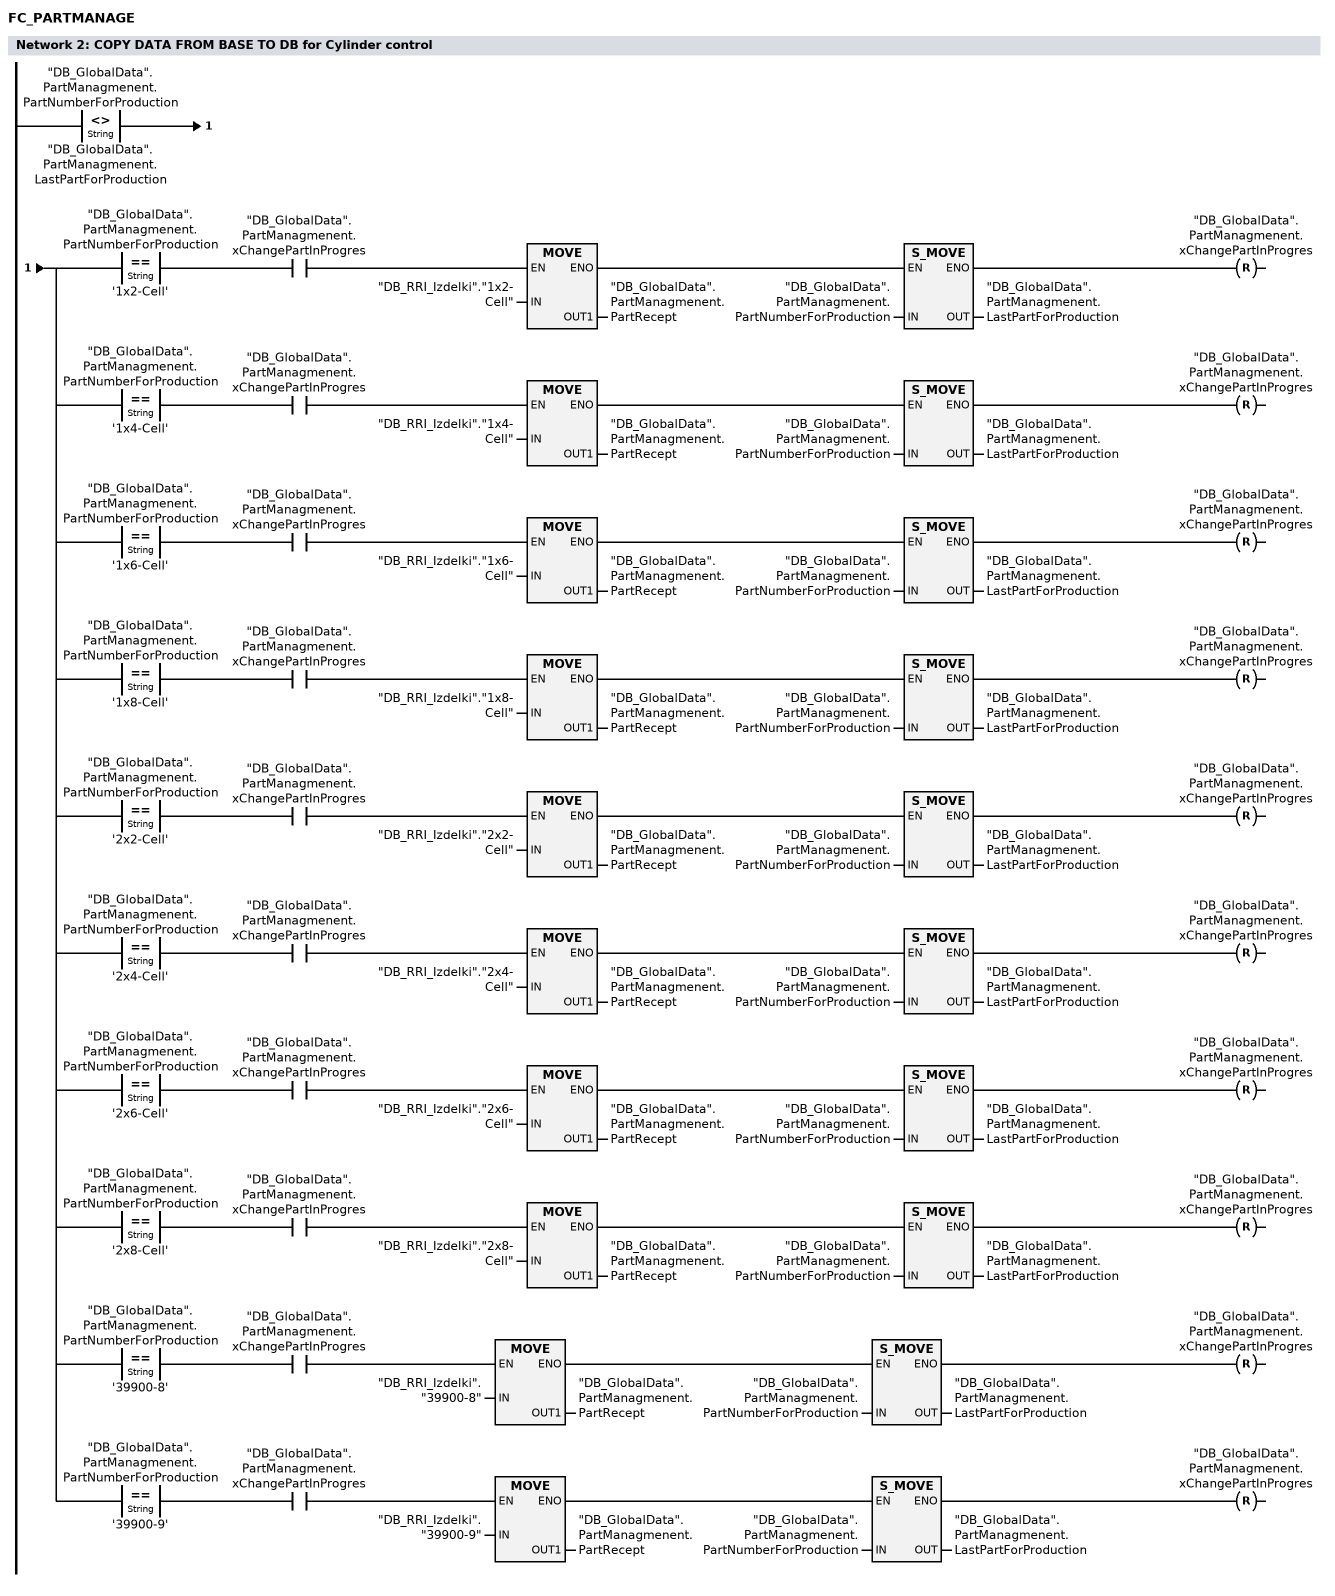
   RUNG wire#powerrail
      { S7_Templates := "SrcType := String" } NE_Contact(in1 := "DB_GlobalData".PartManagmenent.PartNumberForProduction, in2 := "DB_GlobalData".PartManagmenent.LastPartForProduction)
      wire#w1
      { S7_Templates := "SrcType := String" } EQ_Contact(in1 := "DB_GlobalData".PartManagmenent.PartNumberForProduction, in2 := '1x2-Cell')
      Contact( "DB_GlobalData".PartManagmenent.xChangePartInProgres )
      Move(in := "DB_RRI_Izdelki"."1x2-Cell", out1 => "DB_GlobalData".PartManagmenent.PartRecept)
      S_Move(in := "DB_GlobalData".PartManagmenent.PartNumberForProduction, out => "DB_GlobalData".PartManagmenent.LastPartForProduction)
      R_Coil( "DB_GlobalData".PartManagmenent.xChangePartInProgres )
   END_RUNG
   RUNG wire#w1
      { S7_Templates := "SrcType := String" } EQ_Contact(in1 := "DB_GlobalData".PartManagmenent.PartNumberForProduction, in2 := '1x4-Cell')
      Contact( "DB_GlobalData".PartManagmenent.xChangePartInProgres )
      Move(in := "DB_RRI_Izdelki"."1x4-Cell", out1 => "DB_GlobalData".PartManagmenent.PartRecept)
      S_Move(in := "DB_GlobalData".PartManagmenent.PartNumberForProduction, out => "DB_GlobalData".PartManagmenent.LastPartForProduction)
      R_Coil( "DB_GlobalData".PartManagmenent.xChangePartInProgres )
   END_RUNG
   RUNG wire#w1
      { S7_Templates := "SrcType := String" } EQ_Contact(in1 := "DB_GlobalData".PartManagmenent.PartNumberForProduction, in2 := '1x6-Cell')
      Contact( "DB_GlobalData".PartManagmenent.xChangePartInProgres )
      Move(in := "DB_RRI_Izdelki"."1x6-Cell", out1 => "DB_GlobalData".PartManagmenent.PartRecept)
      S_Move(in := "DB_GlobalData".PartManagmenent.PartNumberForProduction, out => "DB_GlobalData".PartManagmenent.LastPartForProduction)
      R_Coil( "DB_GlobalData".PartManagmenent.xChangePartInProgres )
   END_RUNG
   RUNG wire#w1
      { S7_Templates := "SrcType := String" } EQ_Contact(in1 := "DB_GlobalData".PartManagmenent.PartNumberForProduction, in2 := '1x8-Cell')
      Contact( "DB_GlobalData".PartManagmenent.xChangePartInProgres )
      Move(in := "DB_RRI_Izdelki"."1x8-Cell", out1 => "DB_GlobalData".PartManagmenent.PartRecept)
      S_Move(in := "DB_GlobalData".PartManagmenent.PartNumberForProduction, out => "DB_GlobalData".PartManagmenent.LastPartForProduction)
      R_Coil( "DB_GlobalData".PartManagmenent.xChangePartInProgres )
   END_RUNG
   RUNG wire#w1
      { S7_Templates := "SrcType := String" } EQ_Contact(in1 := "DB_GlobalData".PartManagmenent.PartNumberForProduction, in2 := '2x2-Cell')
      Contact( "DB_GlobalData".PartManagmenent.xChangePartInProgres )
      Move(in := "DB_RRI_Izdelki"."2x2-Cell", out1 => "DB_GlobalData".PartManagmenent.PartRecept)
      S_Move(in := "DB_GlobalData".PartManagmenent.PartNumberForProduction, out => "DB_GlobalData".PartManagmenent.LastPartForProduction)
      R_Coil( "DB_GlobalData".PartManagmenent.xChangePartInProgres )
   END_RUNG
   RUNG wire#w1
      { S7_Templates := "SrcType := String" } EQ_Contact(in1 := "DB_GlobalData".PartManagmenent.PartNumberForProduction, in2 := '2x4-Cell')
      Contact( "DB_GlobalData".PartManagmenent.xChangePartInProgres )
      Move(in := "DB_RRI_Izdelki"."2x4-Cell", out1 => "DB_GlobalData".PartManagmenent.PartRecept)
      S_Move(in := "DB_GlobalData".PartManagmenent.PartNumberForProduction, out => "DB_GlobalData".PartManagmenent.LastPartForProduction)
      R_Coil( "DB_GlobalData".PartManagmenent.xChangePartInProgres )
   END_RUNG
   RUNG wire#w1
      { S7_Templates := "SrcType := String" } EQ_Contact(in1 := "DB_GlobalData".PartManagmenent.PartNumberForProduction, in2 := '2x6-Cell')
      Contact( "DB_GlobalData".PartManagmenent.xChangePartInProgres )
      Move(in := "DB_RRI_Izdelki"."2x6-Cell", out1 => "DB_GlobalData".PartManagmenent.PartRecept)
      S_Move(in := "DB_GlobalData".PartManagmenent.PartNumberForProduction, out => "DB_GlobalData".PartManagmenent.LastPartForProduction)
      R_Coil( "DB_GlobalData".PartManagmenent.xChangePartInProgres )
   END_RUNG
   RUNG wire#w1
      { S7_Templates := "SrcType := String" } EQ_Contact(in1 := "DB_GlobalData".PartManagmenent.PartNumberForProduction, in2 := '2x8-Cell')
      Contact( "DB_GlobalData".PartManagmenent.xChangePartInProgres )
      Move(in := "DB_RRI_Izdelki"."2x8-Cell", out1 => "DB_GlobalData".PartManagmenent.PartRecept)
      S_Move(in := "DB_GlobalData".PartManagmenent.PartNumberForProduction, out => "DB_GlobalData".PartManagmenent.LastPartForProduction)
      R_Coil( "DB_GlobalData".PartManagmenent.xChangePartInProgres )
   END_RUNG
   RUNG wire#w1
      { S7_Templates := "SrcType := String" } EQ_Contact(in1 := "DB_GlobalData".PartManagmenent.PartNumberForProduction, in2 := '39900-8')
      Contact( "DB_GlobalData".PartManagmenent.xChangePartInProgres )
      Move(in := "DB_RRI_Izdelki"."39900-8", out1 => "DB_GlobalData".PartManagmenent.PartRecept)
      S_Move(in := "DB_GlobalData".PartManagmenent.PartNumberForProduction, out => "DB_GlobalData".PartManagmenent.LastPartForProduction)
      R_Coil( "DB_GlobalData".PartManagmenent.xChangePartInProgres )
   END_RUNG
   RUNG wire#w1
      { S7_Templates := "SrcType := String" } EQ_Contact(in1 := "DB_GlobalData".PartManagmenent.PartNumberForProduction, in2 := '39900-9')
      Contact( "DB_GlobalData".PartManagmenent.xChangePartInProgres )
      Move(in := "DB_RRI_Izdelki"."39900-9", out1 => "DB_GlobalData".PartManagmenent.PartRecept)
      S_Move(in := "DB_GlobalData".PartManagmenent.PartNumberForProduction, out => "DB_GlobalData".PartManagmenent.LastPartForProduction)
      R_Coil( "DB_GlobalData".PartManagmenent.xChangePartInProgres )
   END_RUNG
   // the same network as SCL:
   #_w1 := "DB_GlobalData".PartManagmenent.PartNumberForProduction <> "DB_GlobalData".PartManagmenent.LastPartForProduction;
   IF #_w1 AND ("DB_GlobalData".PartManagmenent.PartNumberForProduction = '1x2-Cell') AND "DB_GlobalData".PartManagmenent.xChangePartInProgres THEN
       "DB_GlobalData".PartManagmenent.PartRecept := "DB_RRI_Izdelki"."1x2-Cell";
       "DB_GlobalData".PartManagmenent.LastPartForProduction := "DB_GlobalData".PartManagmenent.PartNumberForProduction;
       "DB_GlobalData".PartManagmenent.xChangePartInProgres := FALSE;
   END_IF;
   IF #_w1 AND ("DB_GlobalData".PartManagmenent.PartNumberForProduction = '1x4-Cell') AND "DB_GlobalData".PartManagmenent.xChangePartInProgres THEN
       "DB_GlobalData".PartManagmenent.PartRecept := "DB_RRI_Izdelki"."1x4-Cell";
       "DB_GlobalData".PartManagmenent.LastPartForProduction := "DB_GlobalData".PartManagmenent.PartNumberForProduction;
       "DB_GlobalData".PartManagmenent.xChangePartInProgres := FALSE;
   END_IF;
   IF #_w1 AND ("DB_GlobalData".PartManagmenent.PartNumberForProduction = '1x6-Cell') AND "DB_GlobalData".PartManagmenent.xChangePartInProgres THEN
       "DB_GlobalData".PartManagmenent.PartRecept := "DB_RRI_Izdelki"."1x6-Cell";
       "DB_GlobalData".PartManagmenent.LastPartForProduction := "DB_GlobalData".PartManagmenent.PartNumberForProduction;
       "DB_GlobalData".PartManagmenent.xChangePartInProgres := FALSE;
   END_IF;
   IF #_w1 AND ("DB_GlobalData".PartManagmenent.PartNumberForProduction = '1x8-Cell') AND "DB_GlobalData".PartManagmenent.xChangePartInProgres THEN
       "DB_GlobalData".PartManagmenent.PartRecept := "DB_RRI_Izdelki"."1x8-Cell";
       "DB_GlobalData".PartManagmenent.LastPartForProduction := "DB_GlobalData".PartManagmenent.PartNumberForProduction;
       "DB_GlobalData".PartManagmenent.xChangePartInProgres := FALSE;
   END_IF;
   IF #_w1 AND ("DB_GlobalData".PartManagmenent.PartNumberForProduction = '2x2-Cell') AND "DB_GlobalData".PartManagmenent.xChangePartInProgres THEN
       "DB_GlobalData".PartManagmenent.PartRecept := "DB_RRI_Izdelki"."2x2-Cell";
       "DB_GlobalData".PartManagmenent.LastPartForProduction := "DB_GlobalData".PartManagmenent.PartNumberForProduction;
       "DB_GlobalData".PartManagmenent.xChangePartInProgres := FALSE;
   END_IF;
   IF #_w1 AND ("DB_GlobalData".PartManagmenent.PartNumberForProduction = '2x4-Cell') AND "DB_GlobalData".PartManagmenent.xChangePartInProgres THEN
       "DB_GlobalData".PartManagmenent.PartRecept := "DB_RRI_Izdelki"."2x4-Cell";
       "DB_GlobalData".PartManagmenent.LastPartForProduction := "DB_GlobalData".PartManagmenent.PartNumberForProduction;
       "DB_GlobalData".PartManagmenent.xChangePartInProgres := FALSE;
   END_IF;
   IF #_w1 AND ("DB_GlobalData".PartManagmenent.PartNumberForProduction = '2x6-Cell') AND "DB_GlobalData".PartManagmenent.xChangePartInProgres THEN
       "DB_GlobalData".PartManagmenent.PartRecept := "DB_RRI_Izdelki"."2x6-Cell";
       "DB_GlobalData".PartManagmenent.LastPartForProduction := "DB_GlobalData".PartManagmenent.PartNumberForProduction;
       "DB_GlobalData".PartManagmenent.xChangePartInProgres := FALSE;
   END_IF;
   IF #_w1 AND ("DB_GlobalData".PartManagmenent.PartNumberForProduction = '2x8-Cell') AND "DB_GlobalData".PartManagmenent.xChangePartInProgres THEN
       "DB_GlobalData".PartManagmenent.PartRecept := "DB_RRI_Izdelki"."2x8-Cell";
       "DB_GlobalData".PartManagmenent.LastPartForProduction := "DB_GlobalData".PartManagmenent.PartNumberForProduction;
       "DB_GlobalData".PartManagmenent.xChangePartInProgres := FALSE;
   END_IF;
   IF #_w1 AND ("DB_GlobalData".PartManagmenent.PartNumberForProduction = '39900-8') AND "DB_GlobalData".PartManagmenent.xChangePartInProgres THEN
       "DB_GlobalData".PartManagmenent.PartRecept := "DB_RRI_Izdelki"."39900-8";
       "DB_GlobalData".PartManagmenent.LastPartForProduction := "DB_GlobalData".PartManagmenent.PartNumberForProduction;
       "DB_GlobalData".PartManagmenent.xChangePartInProgres := FALSE;
   END_IF;
   IF #_w1 AND ("DB_GlobalData".PartManagmenent.PartNumberForProduction = '39900-9') AND "DB_GlobalData".PartManagmenent.xChangePartInProgres THEN
       "DB_GlobalData".PartManagmenent.PartRecept := "DB_RRI_Izdelki"."39900-9";
       "DB_GlobalData".PartManagmenent.LastPartForProduction := "DB_GlobalData".PartManagmenent.PartNumberForProduction;
       "DB_GlobalData".PartManagmenent.xChangePartInProgres := FALSE;
   END_IF;
END_REGION
END_FUNCTION

ORGANIZATION_BLOCK "Main"   // OB1, LAD, ProgramCycle
TITLE = "Main Program Sweep (Cycle)"
{ S7_Optimized_Access := 'TRUE' }
VERSION : 0.1
   VAR_INPUT
      Initial_Call : Bool;   // Initial call of this OB
      Remanence : Bool;   // =True, if remanent data are available
   END_VAR
   VAR_TEMP   // added for the SCL form of the ladder/FBD networks
      _w1 : Bool;
      _w2 : Bool;
   END_VAR
BEGIN

REGION Network 1
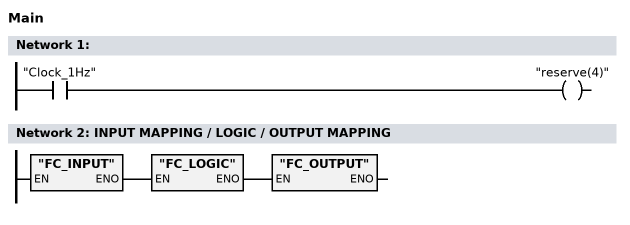
   RUNG wire#powerrail
      Contact( "Clock_1Hz" )
      Coil( "reserve(4)" )
   END_RUNG
   // the same network as SCL:
   "reserve(4)" := "Clock_1Hz";
END_REGION

REGION Network 2: INPUT MAPPING / LOGIC / OUTPUT MAPPING
   RUNG wire#powerrail
      "FC_INPUT"()
      "FC_LOGIC"()
      "FC_OUTPUT"()
   END_RUNG
   // the same network as SCL:
   "FC_INPUT"(ENO => #_w1);
   "FC_LOGIC"(EN := #_w1, ENO => #_w2);
   IF #_w2 THEN "FC_OUTPUT"(); END_IF;
END_REGION
END_ORGANIZATION_BLOCK

// folder: AKD

FUNCTION_BLOCK "FB_AKD"   // FB11, LAD
{ S7_Optimized_Access := 'TRUE' }
VERSION : 0.1
   VAR_INPUT
      bServoEnable : Bool;
      iNastavitevHitrosti : Int;
      dNastavitevPozicije : DInt;
      bPogojiZaVKLOP : Bool;
      iAKD : "AKD_TO_SIEMENS";
      ResetNapake : Bool;
      iStPrograma : Word;
   END_VAR
   VAR_OUTPUT
      oAKD : "SIEMENS_TO_AKD";
      AKDcurrPos : DInt;
      o_BerrStatus : Byte;
      rAKDpos : Real;
      xDriveIsStoped : Bool;
      q_xStartHomming : Bool;
      q_xisHommed : Bool;
      q_xerrNoInTolleranceRange : Bool;
   END_VAR
   VAR_IN_OUT
      iStartHoming : Bool;
      bServoGo : Bool;
   END_VAR
   VAR RETAIN
      TIMER_ON : Array[0..5] of TON_TIME;
   END_VAR
   VAR
      diHitrost : Real;
      dwHitrostRez : Real;
      ServoHommed : Bool;
   END_VAR
   VAR RETAIN
      merker : Array[0..1] of Bool;
   END_VAR
   VAR
      OmogociHome : Bool;
      Varnost : Bool;
      M_varnost : Bool;
      varnostN : Bool;
      TON_fault : TON_TIME;
   END_VAR
   VAR RETAIN
      _xServoGoP : Bool;
      _rCurrntPosition : Real;
      _xServoGoN : Bool;
      _xLastPosition : Real;
   END_VAR
   VAR
      IEC_Timer_0_Instance : TP_TIME;
      R_TRIG_Instance_Home : R_TRIG;
   END_VAR
   VAR RETAIN
      "p_trig-HomePosSet" : Bool;
      "P-trig" : Bool;
      MDI_STATUS : Int;
   END_VAR
   VAR
      statis_target_pos_reach : Bool;
      _errorNotInToleranceRange : Bool;
   END_VAR
   VAR CONSTANT
      AXES_START_MOVING : Int := 10;
      TARGET_POS_REACH : Int := 20;
      RESET_SERVO_GO : Int := 30;
   END_VAR
   VAR_TEMP   // added for the SCL form of the ladder/FBD networks
      _w1 : Bool;
      _w2 : Bool;
      _w3 : Bool;
      _w4 : Bool;
   END_VAR
BEGIN

REGION Network 1: Bool
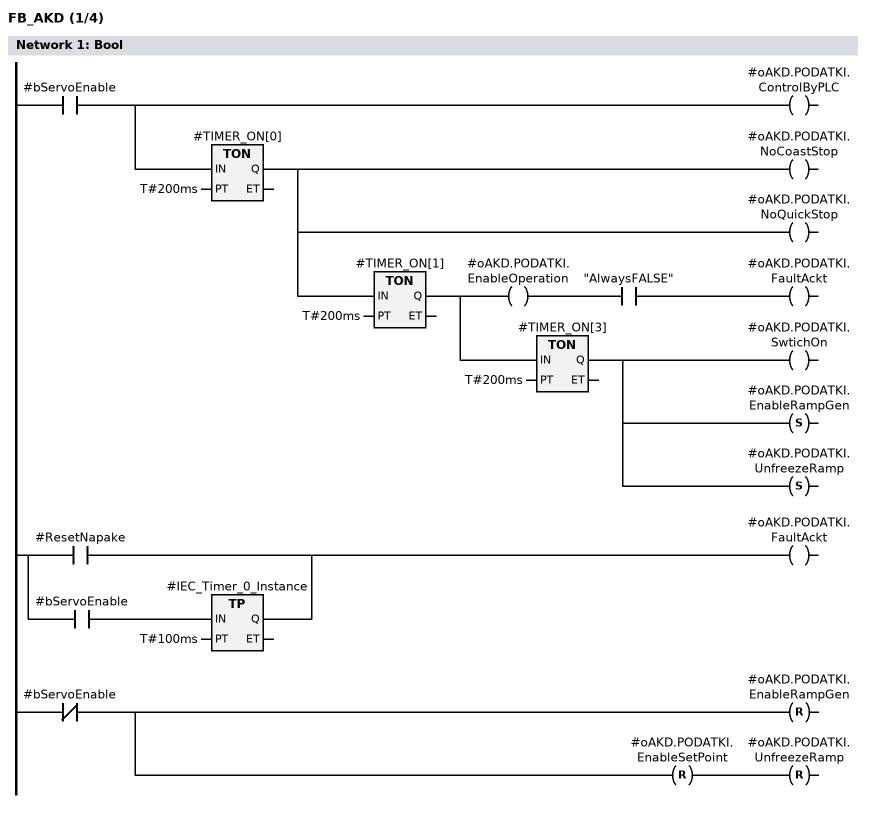
   #oAKD.PODATKI.ControlByPLC := #bServoEnable;
   #TIMER_ON[0].TON(IN := #bServoEnable, PT := T#200ms);
   #oAKD.PODATKI.NoCoastStop := #TIMER_ON[0].Q;
   #oAKD.PODATKI.NoQuickStop := #TIMER_ON[0].Q;
   #TIMER_ON[1].TON(IN := #TIMER_ON[0].Q, PT := T#200ms);
   #oAKD.PODATKI.EnableOperation := #TIMER_ON[1].Q;
   #oAKD.PODATKI.FaultAckt := #TIMER_ON[1].Q AND "AlwaysFALSE";
   #TIMER_ON[3].TON(IN := #TIMER_ON[1].Q, PT := T#200ms);
   #oAKD.PODATKI.SwtichOn := #TIMER_ON[3].Q;
   IF #TIMER_ON[3].Q THEN
       #oAKD.PODATKI.EnableRampGen := TRUE;
       #oAKD.PODATKI.UnfreezeRamp := TRUE;
   END_IF;
   #IEC_Timer_0_Instance(IN := #bServoEnable, PT := T#100ms);   // TP
   #oAKD.PODATKI.FaultAckt := #ResetNapake OR #IEC_Timer_0_Instance.Q;
   IF NOT #bServoEnable THEN
       #oAKD.PODATKI.EnableRampGen := FALSE;
       #oAKD.PODATKI.EnableSetPoint := FALSE;
       #oAKD.PODATKI.UnfreezeRamp := FALSE;
   END_IF;
END_REGION

REGION Network 2: Turn on MDI - manual data inpuit - start task on AKD
   // Requeremnts
   // - S4
   // - mode in position mode (yes)
   // - standard telegram 9 (set at profinet configuration)
   // - axis hommed (homeposset)
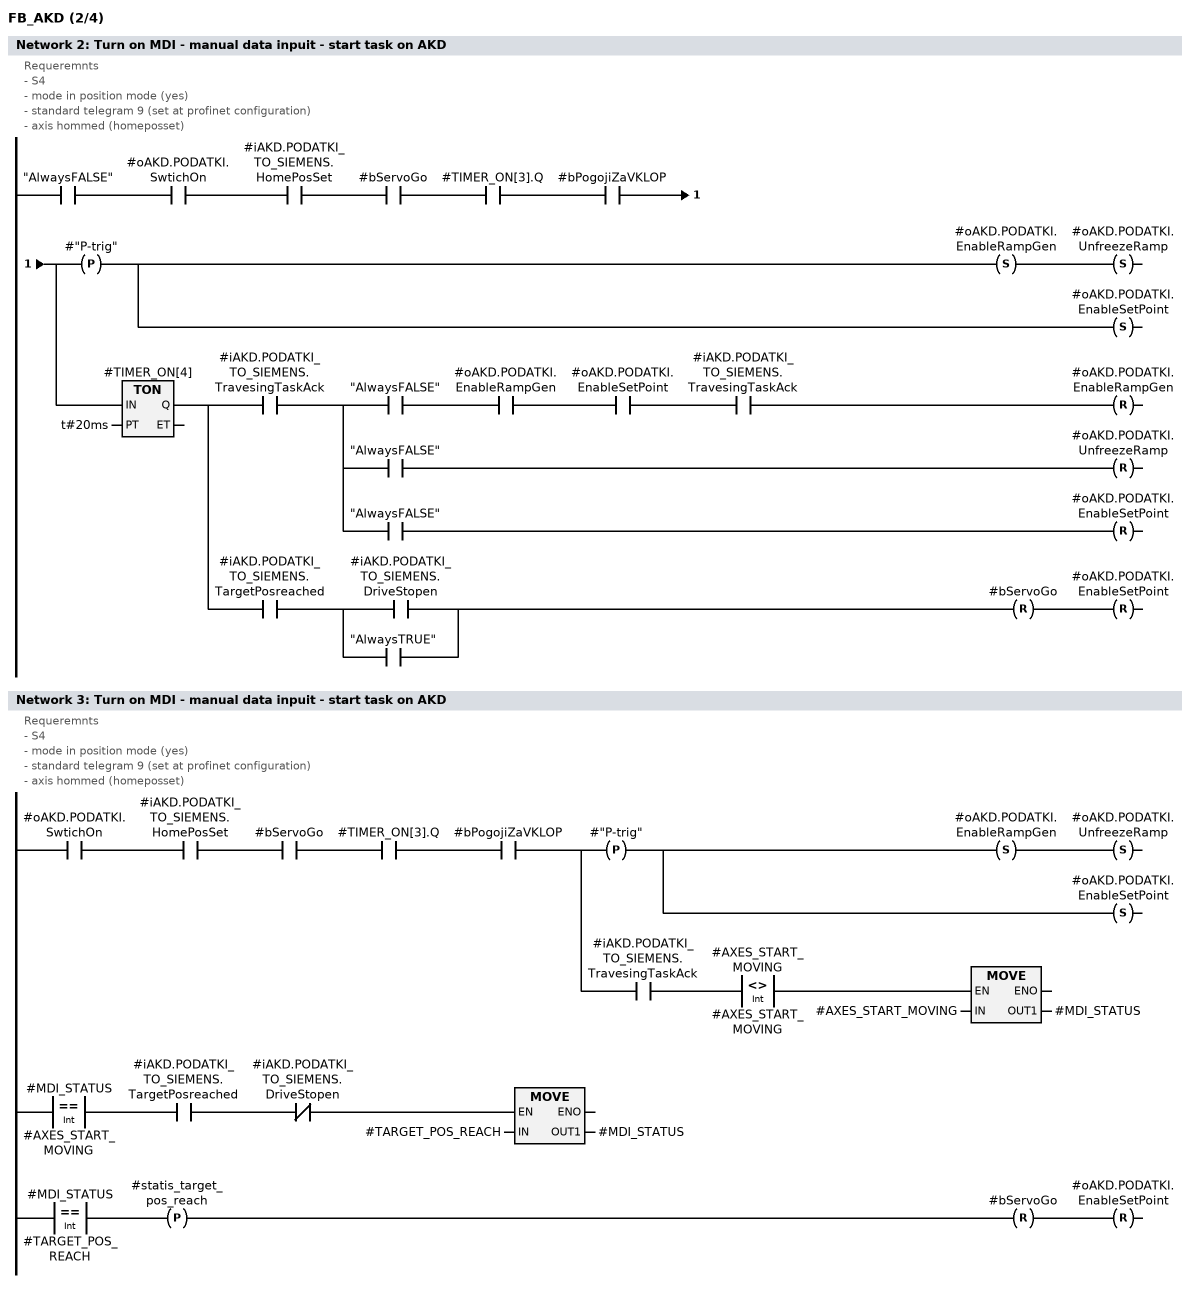
   #_w1 := "AlwaysFALSE" AND #oAKD.PODATKI.SwtichOn AND #iAKD.PODATKI_TO_SIEMENS.HomePosSet AND #bServoGo AND #TIMER_ON[3].Q AND #bPogojiZaVKLOP;
   #_w2 := #_w1 AND NOT #"P-trig";   // rising edge
   #"P-trig" := #_w1;
   IF #_w2 THEN
       #oAKD.PODATKI.EnableRampGen := TRUE;
       #oAKD.PODATKI.UnfreezeRamp := TRUE;
       #oAKD.PODATKI.EnableSetPoint := TRUE;
   END_IF;
   #TIMER_ON[4].TON(IN := #_w1, PT := t#20ms);
   #_w3 := #TIMER_ON[4].Q AND #iAKD.PODATKI_TO_SIEMENS.TravesingTaskAck;
   IF #_w3 AND "AlwaysFALSE" AND #oAKD.PODATKI.EnableRampGen AND #oAKD.PODATKI.EnableSetPoint AND #iAKD.PODATKI_TO_SIEMENS.TravesingTaskAck THEN
       #oAKD.PODATKI.EnableRampGen := FALSE;
   END_IF;
   IF #_w3 AND "AlwaysFALSE" THEN
       #oAKD.PODATKI.UnfreezeRamp := FALSE;
       #oAKD.PODATKI.EnableSetPoint := FALSE;
   END_IF;
   IF #TIMER_ON[4].Q AND #iAKD.PODATKI_TO_SIEMENS.TargetPosreached AND (#iAKD.PODATKI_TO_SIEMENS.DriveStopen OR "AlwaysTRUE") THEN
       #bServoGo := FALSE;
       #oAKD.PODATKI.EnableSetPoint := FALSE;
   END_IF;
END_REGION

REGION Network 3: Turn on MDI - manual data inpuit - start task on AKD
   // Requeremnts
   // - S4
   // - mode in position mode (yes)
   // - standard telegram 9 (set at profinet configuration)
   // - axis hommed (homeposset)
   RUNG wire#powerrail
      Contact( #oAKD.PODATKI.SwtichOn )
      Contact( #iAKD.PODATKI_TO_SIEMENS.HomePosSet )
      Contact( #bServoGo )
      Contact( #TIMER_ON[3].Q )
      Contact( #bPogojiZaVKLOP )
      wire#w1
      P_Trig( #"P-trig" )
      wire#w2
      S_Coil( #oAKD.PODATKI.EnableRampGen )
      S_Coil( #oAKD.PODATKI.UnfreezeRamp )
   END_RUNG
   RUNG wire#w2
      S_Coil( #oAKD.PODATKI.EnableSetPoint )
   END_RUNG
   RUNG wire#w1
      Contact( #iAKD.PODATKI_TO_SIEMENS.TravesingTaskAck )
      { S7_Templates := "SrcType := Int" } NE_Contact(in1 := #AXES_START_MOVING, in2 := #AXES_START_MOVING)
      Move(in := #AXES_START_MOVING, out1 => #MDI_STATUS)
   END_RUNG
   RUNG wire#powerrail
      { S7_Templates := "SrcType := Int" } EQ_Contact(in1 := #MDI_STATUS, in2 := #AXES_START_MOVING)
      Contact( #iAKD.PODATKI_TO_SIEMENS.TargetPosreached )
      I_Contact( #iAKD.PODATKI_TO_SIEMENS.DriveStopen )
      Move(in := #TARGET_POS_REACH, out1 => #MDI_STATUS)
   END_RUNG
   RUNG wire#powerrail
      { S7_Templates := "SrcType := Int" } EQ_Contact(in1 := #MDI_STATUS, in2 := #TARGET_POS_REACH)
      P_Trig( #statis_target_pos_reach )
      R_Coil( #bServoGo )
      R_Coil( #oAKD.PODATKI.EnableSetPoint )
   END_RUNG
   // the same network as SCL:
   #_w1 := #oAKD.PODATKI.SwtichOn AND #iAKD.PODATKI_TO_SIEMENS.HomePosSet AND #bServoGo AND #TIMER_ON[3].Q AND #bPogojiZaVKLOP;
   #_w2 := #_w1 AND NOT #"P-trig";   // rising edge
   #"P-trig" := #_w1;
   IF #_w2 THEN
       #oAKD.PODATKI.EnableRampGen := TRUE;
       #oAKD.PODATKI.UnfreezeRamp := TRUE;
       #oAKD.PODATKI.EnableSetPoint := TRUE;
   END_IF;
   IF #_w1 AND #iAKD.PODATKI_TO_SIEMENS.TravesingTaskAck AND (#AXES_START_MOVING <> #AXES_START_MOVING) THEN
       #MDI_STATUS := #AXES_START_MOVING;
   END_IF;
   IF (#MDI_STATUS = #AXES_START_MOVING) AND #iAKD.PODATKI_TO_SIEMENS.TargetPosreached AND NOT #iAKD.PODATKI_TO_SIEMENS.DriveStopen THEN
       #MDI_STATUS := #TARGET_POS_REACH;
   END_IF;
   #_w3 := #MDI_STATUS = #TARGET_POS_REACH;
   #_w4 := #_w3 AND NOT #statis_target_pos_reach;   // rising edge
   #statis_target_pos_reach := #_w3;
   IF #_w4 THEN
       #bServoGo := FALSE;
       #oAKD.PODATKI.EnableSetPoint := FALSE;
   END_IF;
END_REGION

REGION Network 4
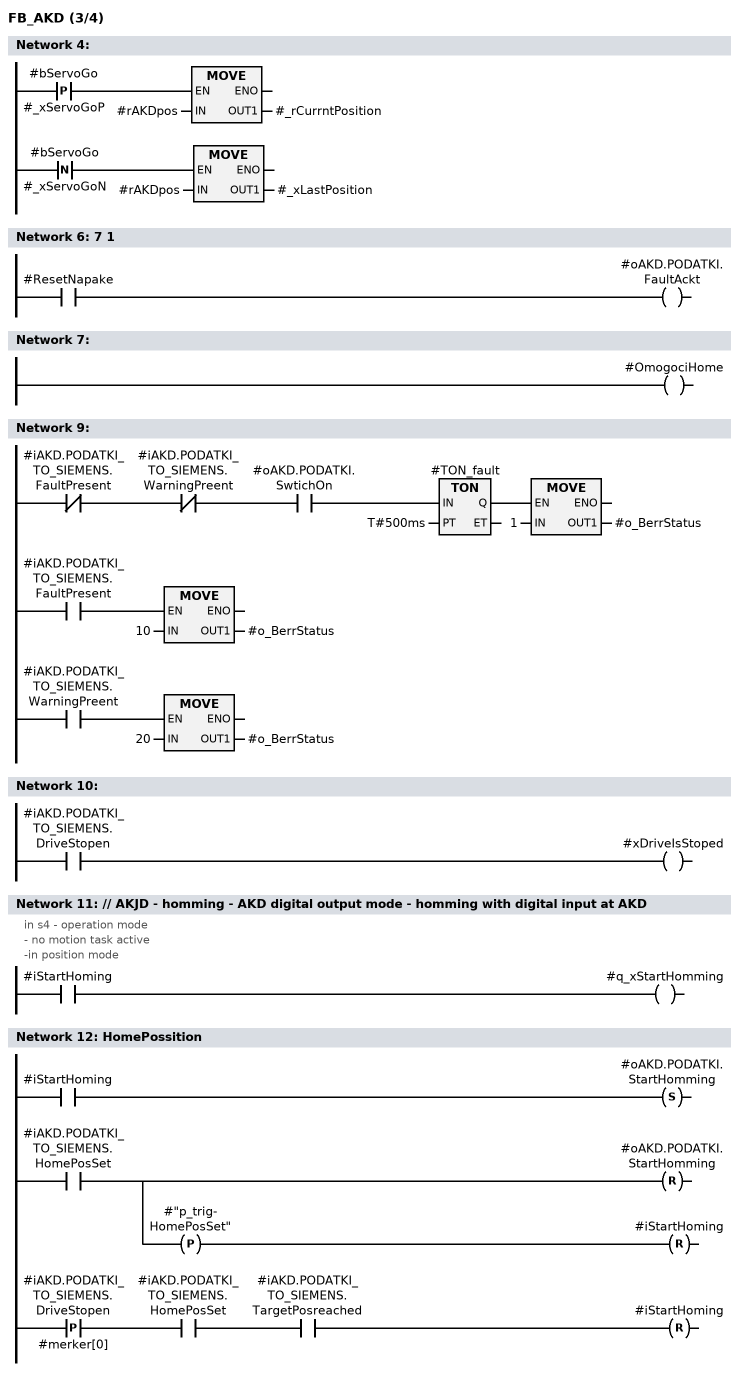
   RUNG wire#powerrail
      P_Contact(operand := #bServoGo, bit := #_xServoGoP)
      Move(in := #rAKDpos, out1 => #_rCurrntPosition)
   END_RUNG
   RUNG wire#powerrail
      N_Contact(operand := #bServoGo, bit := #_xServoGoN)
      Move(in := #rAKDpos, out1 => #_xLastPosition)
   END_RUNG
   // the same network as SCL:
   #_w1 := #bServoGo AND NOT #_xServoGoP;   // rising edge of #bServoGo
   #_xServoGoP := #bServoGo;
   IF #_w1 THEN #_rCurrntPosition := #rAKDpos; END_IF;
   #_w2 := NOT #bServoGo AND #_xServoGoN;   // falling edge of #bServoGo
   #_xServoGoN := #bServoGo;
   IF #_w2 THEN #_xLastPosition := #rAKDpos; END_IF;
END_REGION

REGION Network 5 (SCL)
   //PretvorbaHitrosti
   #diHitrost := INT_TO_REAL(#iNastavitevHitrosti);
   #dwHitrostRez :=((#diHitrost * 4294967295/12000));
   #oAKD.PODATKI.MDI_VELOCITY := REAL_TO_DINT(#dwHitrostRez); //hitrost


   // Operation mode
   #oAKD.PODATKI.MDI_MOD := 16#00_00; //0 - relativni 1//aboslutni gib
   #oAKD.PODATKI.SATANW := #iStPrograma;   //OutputTask

   //pretvorba poziij
   #AKDcurrPos := (#iAKD.PODATKI_TO_SIEMENS.ActualPos * 5 )/ 65536;
   #rAKDpos:= (#iAKD.PODATKI_TO_SIEMENS.ActualPos) / 65536.00;
   //nastavljanjePozicije
   //nastavljanje pozicije
   #oAKD.PODATKI.MDI_TARPOS := (65536 * #dNastavitevPozicije / 5);
END_REGION

REGION Network 6: 7 1
   RUNG wire#powerrail
      Contact( #ResetNapake )
      Coil( #oAKD.PODATKI.FaultAckt )
   END_RUNG
   // the same network as SCL:
   #oAKD.PODATKI.FaultAckt := #ResetNapake;
END_REGION

REGION Network 7
   RUNG wire#powerrail
      Coil( #OmogociHome )
   END_RUNG
   // the same network as SCL:
   #OmogociHome := TRUE;
END_REGION

REGION Network 8: ERROR STATUS
END_REGION

REGION Network 9
   #TON_fault(IN := NOT #iAKD.PODATKI_TO_SIEMENS.FaultPresent AND NOT #iAKD.PODATKI_TO_SIEMENS.WarningPreent AND #oAKD.PODATKI.SwtichOn,   // TON
              PT := T#500ms);
   IF #TON_fault.Q THEN #o_BerrStatus := 1; END_IF;
   IF #iAKD.PODATKI_TO_SIEMENS.FaultPresent THEN #o_BerrStatus := 10; END_IF;
   IF #iAKD.PODATKI_TO_SIEMENS.WarningPreent THEN #o_BerrStatus := 20; END_IF;
END_REGION

REGION Network 10
   RUNG wire#powerrail
      Contact( #iAKD.PODATKI_TO_SIEMENS.DriveStopen )
      Coil( #xDriveIsStoped )
   END_RUNG
   // the same network as SCL:
   #xDriveIsStoped := #iAKD.PODATKI_TO_SIEMENS.DriveStopen;
END_REGION

REGION Network 11: // AKJD - homming - AKD digital output mode - homming with digital input at AKD
   // in s4 - operation mode
   // - no motion task active
   // -in position mode
   RUNG wire#powerrail
      Contact( #iStartHoming )
      Coil( #q_xStartHomming )
   END_RUNG
   // the same network as SCL:
   #q_xStartHomming := #iStartHoming;
END_REGION

REGION Network 12: HomePossition
   RUNG wire#powerrail
      Contact( #iStartHoming )
      S_Coil( #oAKD.PODATKI.StartHomming )
   END_RUNG
   RUNG wire#powerrail
      Contact( #iAKD.PODATKI_TO_SIEMENS.HomePosSet )
      wire#w1
      R_Coil( #oAKD.PODATKI.StartHomming )
   END_RUNG
   RUNG wire#w1
      P_Trig( #"p_trig-HomePosSet" )
      R_Coil( #iStartHoming )
   END_RUNG
   RUNG wire#powerrail
      P_Contact(operand := #iAKD.PODATKI_TO_SIEMENS.DriveStopen, bit := #merker[0])
      Contact( #iAKD.PODATKI_TO_SIEMENS.HomePosSet )
      Contact( #iAKD.PODATKI_TO_SIEMENS.TargetPosreached )
      R_Coil( #iStartHoming )
   END_RUNG
   // the same network as SCL:
   IF #iStartHoming THEN #oAKD.PODATKI.StartHomming := TRUE; END_IF;
   IF #iAKD.PODATKI_TO_SIEMENS.HomePosSet THEN #oAKD.PODATKI.StartHomming := FALSE; END_IF;
   #_w1 := #iAKD.PODATKI_TO_SIEMENS.HomePosSet AND NOT #"p_trig-HomePosSet";   // rising edge
   #"p_trig-HomePosSet" := #iAKD.PODATKI_TO_SIEMENS.HomePosSet;
   IF #_w1 THEN #iStartHoming := FALSE; END_IF;
   #_w2 := #iAKD.PODATKI_TO_SIEMENS.DriveStopen AND NOT #merker[0];   // rising edge of #iAKD.PODATKI_TO_SIEMENS.DriveStopen
   #merker[0] := #iAKD.PODATKI_TO_SIEMENS.DriveStopen;
   IF #_w2 AND #iAKD.PODATKI_TO_SIEMENS.HomePosSet AND #iAKD.PODATKI_TO_SIEMENS.TargetPosreached THEN
       #iStartHoming := FALSE;
   END_IF;
END_REGION

REGION Network 13: OUTPUT : is hommed
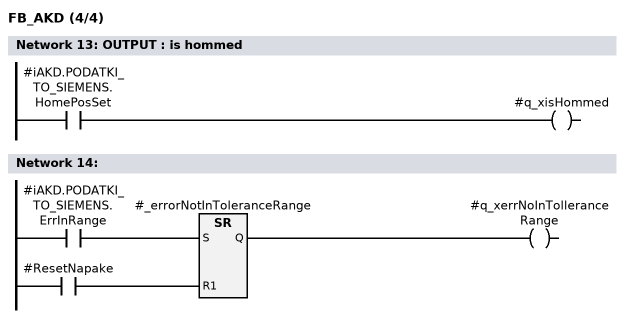
   RUNG wire#powerrail
      Contact( #iAKD.PODATKI_TO_SIEMENS.HomePosSet )
      Coil( #q_xisHommed )
   END_RUNG
   // the same network as SCL:
   #q_xisHommed := #iAKD.PODATKI_TO_SIEMENS.HomePosSet;
END_REGION

REGION Network 14
   RUNG wire#powerrail
      Contact( #iAKD.PODATKI_TO_SIEMENS.ErrInRange )
      S_SR(operand := #_errorNotInToleranceRange, r1 := wire#w1)
      Coil( #q_xerrNoInTolleranceRange )
   END_RUNG
   RUNG wire#powerrail
      Contact( #ResetNapake )
   END_RUNG wire#w1
   // the same network as SCL:
   IF #iAKD.PODATKI_TO_SIEMENS.ErrInRange THEN
       #_errorNotInToleranceRange := TRUE;   // SR flip-flop
   END_IF;
   IF #ResetNapake THEN #_errorNotInToleranceRange := FALSE; END_IF;
   #q_xerrNoInTolleranceRange := #_errorNotInToleranceRange;
END_REGION
END_FUNCTION_BLOCK

FUNCTION_BLOCK "AKD_PN_TG400_v05"   // FB14, SCL
TITLE = AKD_PN_TG400_TIA13_v05
{ S7_Optimized_Access := 'FALSE' }
AUTHOR : jcoleman
FAMILY : TG400
VERSION : 5.0
// This function block supports Profinet communication with the AKD drive using Telegram 400.  It is written in TIA V13. 
// For more information, please see the AKD Profinet Manual and the supporting documentation for this function block.
   VAR_INPUT
      iID : Hw_Io;   // Hardware identifier
      iInit : Bool;   // initialize config for TG400
      iEStop : Bool;   // immediate quick stop and disable
      iSW_Enable : Bool;   // enable/disable
      iStop : Bool;   // stop all movement
      iReset : Bool;   // reset drive faults
      iStart_Homing : Bool;   // start homing
      iStart_Jog : Bool;   // start jog
      iStart_Move : Bool;   // start motion task
      iMT_Pause : Bool;   // pause active motion task
      iMT_MoveType : Word;   // motion task control word 0 = relative; 1 = absolute
      iMTNum : Word;   // motion task number 0x8000 = direct motion task
      iCmdPos : DWord;   // commanded position for motion task or homing
      iCmdVel : DWord;   // commanded velocity for jog or direct motion task
      iCmdAcc : Word;   // commanded acceleration for jog or direct motion task
      iCmdDec : Word;   // commanded deceleration for jog or direct motion task
   END_VAR
   VAR_OUTPUT
      oInitDone : Bool;   // initialization status - 0 while configuring TG400, 1= done
      oStatus : DWord;   // ZSW1
      oPos : DWord;   // actual position
      oVel : Word;   // actual velocity x * 12000 rpm / 2^15
      oCurrent : Word;   // actual current x *DRV.IPEAK / 2^14
      oEnabled : Bool;   // Drive power on
      oError : Bool;   // fault in function block or communication
      oMoving : Bool;   // axis enabled and moving
      oHomed : Bool;   // axis homed
      oInPos : Bool;   // axis within in-position window
      oFault : Bool;   // drive fault
      oWarning : Bool;   // drive warning
   END_VAR
   VAR
      TG_400 : "UDT_AKD_TG400";
      wPNReadStatus : Word;
      bPNReadError : Bool;
      wPNWriteStatus : Word;
      bPNWriteError : Bool;
      bResetDone : Bool;
      bHomeStarted : Bool;
      bStartMoveDone : Bool;
      bEstop : Bool;
      wStartReset : Int;
      wStartMove : Int;
      wSDOStatus : Word;
      bySDODataArray : Array[0..63] of Byte;
      SDOWrite : WRREC;
      SDORead : RDREC;
      bSDOReq : Bool;
      bSDOWriteBusy : Bool;
      bSDOWriteDone : Bool;
      bSDOWriteError : Bool;
      bSDOReadBusy : Bool;
      bSDOReadDone : Bool;
      bSDOReadError : Bool;
      wSDOReadValue : Word;
      wSDOAddress : Word;
      bSWEnabled : Bool;
      wHomingStartPoint : Word;
      bStartMove : Bool;
      bSDOStatusReadActive : Bool;
   END_VAR
BEGIN
   ////////////////////////////////////////////////////////////////////////////////////////////////////////
   // Standard communication module between a Kollmorgen AKD and S7-1200/1500 PLC
   //
   // Version  When        Who         What
   // ---------------------------------------------
   // V 05     09.05.17    JColeman KM Changed Telegram 400 mapping PNU writes to be individual writes, rather
   //                                  than a block write...to be more robust.
   // V 04     08.31.17    JColeman KM Changed error handling to indicate internal block errors.
   // V 03     06.05.17    JColeman KM Changed EStop code to set flag without waiting for motion to stop. 
   //                                  Added setting opmode=2 in init section.
   //                                  Added comments.
   //                                  Added information to FB properties.
   //                                  Turn on real-time jog mode during enable process.
   //                                  Do not use Optimized block access.
   // V 02     05.12.17    JColeman KM Changed names of inputs and outputs to be more user friendly
   //                                  Added output oInitDone to indicate when the telegram configuration is complete
   //                                  Changed name of FB to be specific to TG400
   //                                  Changed verion numbering
   // V 1.000  17.09.15    MRupf KM    Conversion to TIA V13 SP1
   // V 0.004  09.07.15    MRupf KM    Home_dist changed to DINT variable length
   //          06.07.15    MRupf KM    Fault and Warning read locked angainst interruption
   // V 0.003  05.06.15    MRupf KM    New iStart_MT is only accepted after the ZSW1 Bit 12 is FALSE again
   //          03.06.15    MRupf KM    Handshake to start motion task with ZSW1 Bit 12 and auto reset after 500ms #285
   //          14.04.15    MRupf KM    Init write cases extended to not do endless recall on error
   //                                  Homing start stop bug, #246-250
   //                                  Reset STW1.6/.7 only after two PN cylce #214, 283
   // V 0.002  26.02.15    MRupf KM    Setup Telegramm 400 with HOME.DIST, VL.FB, IL.FB
   //                                  Read Fault and Warning No. if acitve
   //                                  Reset STW if drive fault happens while enabled    
   // V 0.001  18.02.15    MRupf KM    First version
   //////////////////////////////////////////////////////////////////////////////////////////////////////////

   // initialisation
   IF #iInit THEN
       #wSDOStatus := 0;
       #oInitDone := FALSE;    //False during telegram configuration
   END_IF;
   IF #wSDOStatus < 20 THEN //set telegram send data = 0
       #TG_400.Send.STW1 := 0;
       #TG_400.Send.SATZANW := 0;
       #TG_400.Send.STW2 := 0;
       #TG_400.Send.MDI_TARPOS := 0;
       #TG_400.Send.MDI_VELOCITY := 0;
       #TG_400.Send.MDI_ACC := 0;
       #TG_400.Send.MDI_DEC := 0;
       #TG_400.Send.MDI_MOD := 0;

       #bPNReadError := FALSE;
       #bPNWriteError := FALSE;
   END_IF;

   // Do the setup of the Telegram 400
   IF NOT #iInit AND #wSDOStatus < 19 THEN

       // Map Telegram 400 Send
       // Clear the Array and start the request
       IF #wSDOStatus = 0 THEN
           FILL_BLK(IN := 0,
                    COUNT := 64,
                    OUT => #bySDODataArray[0]);
           #bSDOReq := TRUE;
           #bSDOWriteDone := FALSE;
           #wSDOStatus := 1; //proceed to Step 1
       END_IF;
       // setup the array data and start WRREC
       IF #wSDOStatus = 1 THEN //Step 1
           #bySDODataArray[0] := 16#ff; //Request Reference
           #bySDODataArray[1] := 16#02; //2 for write PNU
           #bySDODataArray[2] := 16#00; //Axis# is 0 for AKD
           #bySDODataArray[3] := 16#01; //number of parameters
           // Set PNU 915 subindex 8
           #bySDODataArray[4] := 16#10; //Attribute is 0x10
           #bySDODataArray[5] := 16#01; //Number of elements =1
           #bySDODataArray[6] := 16#03; //0x393 for PNU 915
           #bySDODataArray[7] := 16#93; //PNU 915
           #bySDODataArray[8] := 16#00; //subindex
           #bySDODataArray[9] := 16#08; //subindex 8 for 8th word of telegram
           // To PNU 100 (HOME.DIST)
           #bySDODataArray[10] := 16#42; //Format =0x42 for Word
           #bySDODataArray[11] := 16#01; //Number of values
           #bySDODataArray[12] := 16#00; //data
           #bySDODataArray[13] := 16#64; //data - Signal #100 for HOME.DIST

           #SDOWrite(REQ := #bSDOReq, //do the PNU write
                     ID := #iID,
                     INDEX := 47, //AKD suppors "Record Data 47"
                     LEN := 14,   //data length
                     BUSY => #bSDOWriteBusy,
                     DONE => #bSDOWriteDone,
                     ERROR => #bSDOWriteError,
                     RECORD := #bySDODataArray);
           IF #bSDOWriteBusy THEN
               #bSDOReq := FALSE;
           ELSIF #bSDOWriteDone THEN
               #wSDOStatus := 2; //proceed to Step 2
           END_IF;
       END_IF;

       // Map Telegram 400 Receive
       // Clear the Array and start the request
       IF #wSDOStatus = 2 THEN //Step 2
           FILL_BLK(IN := 0,
                    COUNT := 64,
                    OUT => #bySDODataArray[0]);
           #bSDOReq := TRUE;
           #bSDOWriteDone := FALSE;
           #wSDOStatus := 3; //proceed to Step 3
       END_IF;
       // setup the array data and start WRREC
       IF #wSDOStatus = 3 THEN //Step 3
           #bySDODataArray[0] := 16#fe; //Request Reference
           #bySDODataArray[1] := 16#02; //2 for write PNU
           #bySDODataArray[2] := 16#00; //Axis# is 0 for AKD
           #bySDODataArray[3] := 16#01; // Number of parameters to write at a time
           // Set PNU 916 subindex 0
           #bySDODataArray[4] := 16#10; //Attribute is 0x10
           #bySDODataArray[5] := 16#01; //Number of elements =1
           #bySDODataArray[6] := 16#03; //0x394 for PNU 916
           #bySDODataArray[7] := 16#94; //PNU 916
           #bySDODataArray[8] := 16#00; //subindex
           #bySDODataArray[9] := 16#00; //subindex 0 for 1st word of telegram
           // To PNU 2 (ZSW1)
           #bySDODataArray[10] := 16#42; //Format =0x42 for Word
           #bySDODataArray[11] := 16#01; //Number of values
           #bySDODataArray[12] := 16#00; //data
           #bySDODataArray[13] := 16#02; //data - Signal #2 (0x02) for ZSW1

           #SDOWrite(REQ := #bSDOReq, //do the PNU write
                     ID := #iID,
                     INDEX := 47, //AKD suppors "Record Data 47"
                     LEN := 14,   //data length
                     BUSY => #bSDOWriteBusy,
                     DONE => #bSDOWriteDone,
                     ERROR => #bSDOWriteError,
                     RECORD := #bySDODataArray);
           IF #bSDOWriteBusy THEN
               #bSDOReq := FALSE;
           ELSIF #bSDOWriteDone THEN
               #wSDOStatus := 4; //proceed to Step 4
           END_IF;
       END_IF;

       // Clear the Array and start the request
       IF #wSDOStatus = 4 THEN //Step 4
           FILL_BLK(IN := 0,
                    COUNT := 64,
                    OUT => #bySDODataArray[0]);
           #bSDOReq := TRUE;
           #bSDOWriteDone := FALSE;
           #wSDOStatus := 5; //proceed to Step 5
       END_IF;
       // setup the array data and start WRREC
       IF #wSDOStatus = 5 THEN //Step 5
           #bySDODataArray[0] := 16#fd; //Request Reference
           #bySDODataArray[1] := 16#02; //2 for write PNU
           #bySDODataArray[2] := 16#00; //Axis# is 0 for AKD
           #bySDODataArray[3] := 16#01; // Number of parameters to write at a time
           // Set PNU 916 subindex 1
           #bySDODataArray[4] := 16#10; //Attribute is 0x10
           #bySDODataArray[5] := 16#01; //Number of elements =1
           #bySDODataArray[6] := 16#03; //0x394 for PNU 916
           #bySDODataArray[7] := 16#94; //PNU 916
           #bySDODataArray[8] := 16#00; //subindex
           #bySDODataArray[9] := 16#01; //subindex 1 for 2nd word of telegram
           // To PNU 33 (AKTSATZ)
           #bySDODataArray[10] := 16#42; //Format =0x42 for Word
           #bySDODataArray[11] := 16#01; //Number of values
           #bySDODataArray[12] := 16#00; //data
           #bySDODataArray[13] := 16#21; //data - Signal #33 (0x21) for AKTSATZ

           #SDOWrite(REQ := #bSDOReq, //do the PNU write
                     ID := #iID,
                     INDEX := 47, //AKD suppors "Record Data 47"
                     LEN := 14,   //data length
                     BUSY => #bSDOWriteBusy,
                     DONE => #bSDOWriteDone,
                     ERROR => #bSDOWriteError,
                     RECORD := #bySDODataArray);
           IF #bSDOWriteBusy THEN
               #bSDOReq := FALSE;
           ELSIF #bSDOWriteDone THEN
               #wSDOStatus := 6; //proceed to Step 6
           END_IF;
       END_IF;

       // Clear the Array and start the request
       IF #wSDOStatus = 6 THEN //Step 6
           FILL_BLK(IN := 0,
                    COUNT := 64,
                    OUT => #bySDODataArray[0]);
           #bSDOReq := TRUE;
           #bSDOWriteDone := FALSE;
           #wSDOStatus := 7; //proceed to Step 7
       END_IF;
       // setup the array data and start WRREC
       IF #wSDOStatus = 7 THEN //Step 7
           #bySDODataArray[0] := 16#fc; //Request Reference
           #bySDODataArray[1] := 16#02; //2 for write PNU
           #bySDODataArray[2] := 16#00; //Axis# is 0 for AKD
           #bySDODataArray[3] := 16#01; // Number of parameters to write at a time
           // Set PNU 916 subindex 2
           #bySDODataArray[4] := 16#10; //Attribute is 0x10
           #bySDODataArray[5] := 16#01; //Number of elements =1
           #bySDODataArray[6] := 16#03; //0x394 for PNU 916
           #bySDODataArray[7] := 16#94; //PNU 916
           #bySDODataArray[8] := 16#00; //subindex
           #bySDODataArray[9] := 16#02; //subindex 2 for 3rd word of telegram
           // To PNU 4 (ZSW1)
           #bySDODataArray[10] := 16#42; //Format =0x42 for Word
           #bySDODataArray[11] := 16#01; //Number of values
           #bySDODataArray[12] := 16#00; //data
           #bySDODataArray[13] := 16#04; //data - Signal #4 (0x04) for ZSW2

           #SDOWrite(REQ := #bSDOReq, //do the PNU write
                     ID := #iID,
                     INDEX := 47, //AKD suppors "Record Data 47"
                     LEN := 14,   //data length
                     BUSY => #bSDOWriteBusy,
                     DONE => #bSDOWriteDone,
                     ERROR => #bSDOWriteError,
                     RECORD := #bySDODataArray);
           IF #bSDOWriteBusy THEN
               #bSDOReq := FALSE;
           ELSIF #bSDOWriteDone THEN
               #wSDOStatus := 8; //proceed to Step 8
           END_IF;
       END_IF;

       // Clear the Array and start the request
       IF #wSDOStatus = 8 THEN //Step 8
           FILL_BLK(IN := 0,
                    COUNT := 64,
                    OUT => #bySDODataArray[0]);
           #bSDOReq := TRUE;
           #bSDOWriteDone := FALSE;
           #wSDOStatus := 9; //proceed to Step 9
       END_IF;
       // setup the array data and start WRREC
       IF #wSDOStatus = 9 THEN //Step 9
           #bySDODataArray[0] := 16#fb; //Request Reference
           #bySDODataArray[1] := 16#02; //2 for write PNU
           #bySDODataArray[2] := 16#00; //Axis# is 0 for AKD
           #bySDODataArray[3] := 16#01; // Number of parameters to write at a time
           // Set PNU 916 subindex 3
           #bySDODataArray[4] := 16#10; //Attribute is 0x10
           #bySDODataArray[5] := 16#01; //Number of elements =1
           #bySDODataArray[6] := 16#03; //0x394 for PNU 916
           #bySDODataArray[7] := 16#94; //PNU 916
           #bySDODataArray[8] := 16#00; //subindex
           #bySDODataArray[9] := 16#03; //subindex 3 for 4th word of telegram
           // To PNU 28 (XIST_A)
           #bySDODataArray[10] := 16#42; //Format =0x42 for Word
           #bySDODataArray[11] := 16#01; //Number of values
           #bySDODataArray[12] := 16#00; //data
           #bySDODataArray[13] := 16#1C; //data - Signal #28 (0x1C) for XIST_A

           #SDOWrite(REQ := #bSDOReq, //do the PNU write
                     ID := #iID,
                     INDEX := 47, //AKD suppors "Record Data 47"
                     LEN := 14,   //data length
                     BUSY => #bSDOWriteBusy,
                     DONE => #bSDOWriteDone,
                     ERROR => #bSDOWriteError,
                     RECORD := #bySDODataArray);
           IF #bSDOWriteBusy THEN
               #bSDOReq := FALSE;
           ELSIF #bSDOWriteDone THEN
               #wSDOStatus := 10; //proceed to Step 10
           END_IF;
       END_IF;

       // Clear the Array and start the request
       IF #wSDOStatus = 10 THEN //Step 10
           FILL_BLK(IN := 0,
                    COUNT := 64,
                    OUT => #bySDODataArray[0]);
           #bSDOReq := TRUE;
           #bSDOWriteDone := FALSE;
           #wSDOStatus := 11; //proceed to Step 11
       END_IF;
       // setup the array data and start WRREC
       IF #wSDOStatus = 11 THEN //Step 11
           #bySDODataArray[0] := 16#fa; //Request Reference
           #bySDODataArray[1] := 16#02; //2 for write PNU
           #bySDODataArray[2] := 16#00; //Axis# is 0 for AKD
           #bySDODataArray[3] := 16#01; // Number of parameters to write at a time
           // Set PNU 916 subindex 4
           #bySDODataArray[4] := 16#10; //Attribute is 0x10
           #bySDODataArray[5] := 16#01; //Number of elements =1
           #bySDODataArray[6] := 16#03; //0x394 for PNU 916
           #bySDODataArray[7] := 16#94; //PNU 916
           #bySDODataArray[8] := 16#00; //subindex
           #bySDODataArray[9] := 16#04; //subindex 4 for 5th word of telegram
           // To PNU 6 (NIST_A)
           #bySDODataArray[10] := 16#42; //Format =0x42 for Word
           #bySDODataArray[11] := 16#01; //Number of values
           #bySDODataArray[12] := 16#00; //data
           #bySDODataArray[13] := 16#06; //data - Signal #6 (0x06) for NIST_A (VL.FB)

           #SDOWrite(REQ := #bSDOReq, //do the PNU write
                     ID := #iID,
                     INDEX := 47, //AKD suppors "Record Data 47"
                     LEN := 14,   //data length
                     BUSY => #bSDOWriteBusy,
                     DONE => #bSDOWriteDone,
                     ERROR => #bSDOWriteError,
                     RECORD := #bySDODataArray);
           IF #bSDOWriteBusy THEN
               #bSDOReq := FALSE;
           ELSIF #bSDOWriteDone THEN
               #wSDOStatus := 12; //proceed to Step 12
           END_IF;
       END_IF;